screen "Error Counter_2" 320x240
   TextField "Text field_1" at 26,1 size 269x18; Text 'CURRENT SHIFT DATA MINUS 2 (Detil Error)'
   Button "Button_3" at 6,199 size 45x34; TextOff 'Main Page'; PictureOff "Home"
      on Click: ActivateScreen("Main Page", 0)
   Button "Button_1" at 57,206 size 93x28; TextOff 'Back To Data Statistika'; TextOn 'Data Statistika'
      on Click: ActivateScreen("Data Statistika", 0)
   Button "Button_2" at 206,206 size 97x28; TextOff '<----- Back'; TextOn 'Sloft Data'
      on Click: ActivateScreen("Data Time Current Shift_2", 0)
   IOField "I/O field_6" at 6,19 size 132x18; FormatPattern 9999999999999999999999999999999999999999
      ProcessValue <- "DB_DTL1_Cur_ShiftA_2"
   TextField "Text field_9" at 145,21 size 19x15; Text 'S/D'
   IOField "I/O field_7" at 169,20 size 132x18; FormatPattern 9999999999999999999999999999999999999999
      ProcessValue <- "DB_DTL1_Cur_ShiftB_2"
   TextField "Text field_34" at 6,153 size 21x19; Text '6'
   TextField "Text field_33" at 7,133 size 21x19; Text '5'
   TextField "Text field_32" at 7,114 size 21x19; Text '4'
   TextField "Text field_31" at 7,95 size 21x19; Text '3'
   TextField "Text field_30" at 7,76 size 21x19; Text '2'
   TextField "Text field_29" at 7,58 size 21x19; Text '1'
   TextField "Text field_28" at 7,40 size 21x19; Text 'No'
   IOField "I/O field_8" at 225,153 size 26x19; FormatPattern 999
      ProcessValue <- "DB_DTLData_DTL_RS Pneu Er_2.SECOND"
   IOField "I/O field_16" at 200,153 size 25x19; FormatPattern 999
      ProcessValue <- "DB_DTLData_DTL_RS Pneu Er_2.MINUTE"
   IOField "I/O field_17" at 175,153 size 25x19; FormatPattern 999
      ProcessValue <- "DB_DTLData_DTL_RS Pneu Er_2.HOUR"
   TextField "Text field_8" at 29,153 size 145x19; Text 'Reed Swicth Pneumatic Error'
   TextField "Text field_10" at 196,152 size 8x17; Text ':'
   TextField "Text field_21" at 220,153 size 8x17; Text ':'
   IOField "I/O field_21" at 225,94 size 26x19; FormatPattern 999
      ProcessValue <- "Data_DTLData_DTL_Imaje Not In Position[2].SECOND"
   IOField "I/O field_22" at 200,94 size 25x19; FormatPattern 999
      ProcessValue <- "Data_DTLData_DTL_Imaje Not In Position[2].MINUTE"
   IOField "I/O field_23" at 175,94 size 25x19; FormatPattern 999
      ProcessValue <- "Data_DTLData_DTL_Imaje Not In Position[2].HOUR"
   TextField "Text field_25" at 29,95 size 145x19; Text 'Imaje Not In Position'
   IOField "I/O field_18" at 225,76 size 26x19; FormatPattern 999
      ProcessValue <- "Data_DTLData_DTL_Paper R Out[2].SECOND"
   IOField "I/O field_19" at 200,76 size 25x19; FormatPattern 999
      ProcessValue <- "Data_DTLData_DTL_Paper R Out[2].MINUTE"
   IOField "I/O field_20" at 175,76 size 25x19; FormatPattern 999
      ProcessValue <- "Data_DTLData_DTL_Paper R Out[2].HOUR"
   TextField "Text field_22" at 29,76 size 145x19; Text 'Imaje Papper Or Ribbon Out'
   TextField "Text field_2" at 176,43 size 24x15; Text 'Hour'
   IOField "I/O field_10" at 225,134 size 26x19; FormatPattern 999
      ProcessValue <- "DB_DTLData_DTL_Slof Jam_2.SECOND"
   IOField "I/O field_11" at 200,134 size 25x19; FormatPattern 999
      ProcessValue <- "DB_DTLData_DTL_Slof Jam_2.MINUTE"
   IOField "I/O field_12" at 175,134 size 25x19; FormatPattern 999
      ProcessValue <- "DB_DTLData_DTL_Slof Jam_2.HOUR"
   IOField "I/O field_4" at 225,114 size 26x19; FormatPattern 999
      ProcessValue <- "DB_DTLData_DTL_Press Low_2.SECOND"
   IOField "I/O field_5" at 200,114 size 25x19; FormatPattern 999
      ProcessValue <- "DB_DTLData_DTL_Press Low_2.MINUTE"
   IOField "I/O field_9" at 175,114 size 25x19; FormatPattern 999
      ProcessValue <- "DB_DTLData_DTL_Press Low_2.HOUR"
   TextField "Text field_12" at 229,43 size 19x15; Text 'Sec'
   TextField "Text field_11" at 203,43 size 19x15; Text 'Min'
   IOField "I/O field_2" at 225,59 size 26x19; FormatPattern 999
      ProcessValue <- "DB_DTLData_DTL_Imaje Er_2.SECOND"
   IOField "I/O field_1" at 200,59 size 25x19; FormatPattern 999
      ProcessValue <- "DB_DTLData_DTL_Imaje Er_2.MINUTE"
   TextField "Text field_3" at 30,42 size 144x17; Text 'Error Counter'
   TextField "Text field_4" at 29,59 size 145x19; Text 'System Imaje Error'
   TextField "Text field_5" at 29,114 size 145x21; Text 'Pressure Low'
   TextField "Text field_6" at 29,133 size 145x20; Text 'Sloft Jammed'
   IOField "I/O field_3" at 175,59 size 25x19; FormatPattern 999
      ProcessValue <- "DB_DTLData_DTL_Imaje Er_2.HOUR"
   TextField "Text field_13" at 196,58 size 8x17; Text ':'
   TextField "Text field_14" at 196,113 size 8x17; Text ':'
   TextField "Text field_15" at 196,133 size 8x17; Text ':'
   TextField "Text field_17" at 220,58 size 8x17; Text ':'
   TextField "Text field_18" at 220,113 size 8x17; Text ':'
   TextField "Text field_19" at 220,133 size 8x17; Text ':'
   TextField "Text field_23" at 196,75 size 8x17; Text ':'
   TextField "Text field_24" at 220,75 size 8x17; Text ':'
   TextField "Text field_26" at 196,93 size 8x17; Text ':'
   TextField "Text field_27" at 220,93 size 8x17; Text ':'

screen "Error Counter_3" 320x240
   TextField "Text field_1" at 24,1 size 269x18; Text 'CURRENT SHIFT DATA MINUS 3 (Detil Error)'
   Button "Button_3" at 3,198 size 45x34; TextOff 'Main Page'; PictureOff "Home"
      on Click: ActivateScreen("Main Page", 0)
   Button "Button_1" at 54,203 size 93x28; TextOff 'Back To Data Statistika'; TextOn 'Data Statistika'
      on Click: ActivateScreen("Data Statistika", 0)
   Button "Button_2" at 206,203 size 97x28; TextOff '<----- Back'; TextOn 'Sloft Data'
      on Click: ActivateScreen("Data Time Current Shift_3", 0)
   IOField "I/O field_6" at 6,20 size 132x18; FormatPattern 9999999999999999999999999999999999999999
      ProcessValue <- "DB_DTL1_Cur_ShiftA_3"
   TextField "Text field_9" at 145,24 size 19x15; Text 'S/D'
   IOField "I/O field_7" at 169,21 size 132x18; FormatPattern 9999999999999999999999999999999999999999
      ProcessValue <- "DB_DTL1_Cur_ShiftB_3"
   TextField "Text field_34" at 6,153 size 21x19; Text '6'
   TextField "Text field_33" at 7,133 size 21x19; Text '5'
   TextField "Text field_32" at 7,114 size 21x19; Text '4'
   TextField "Text field_31" at 7,95 size 21x19; Text '3'
   TextField "Text field_30" at 7,76 size 21x19; Text '2'
   TextField "Text field_29" at 7,58 size 21x19; Text '1'
   TextField "Text field_28" at 7,40 size 21x19; Text 'No'
   IOField "I/O field_8" at 225,153 size 26x19; FormatPattern 999
      ProcessValue <- "DB_DTLData_DTL_RS Pneu Er_3.SECOND"
   IOField "I/O field_16" at 200,153 size 25x19; FormatPattern 999
      ProcessValue <- "DB_DTLData_DTL_RS Pneu Er_3.MINUTE"
   IOField "I/O field_17" at 175,153 size 25x19; FormatPattern 999
      ProcessValue <- "DB_DTLData_DTL_RS Pneu Er_3.HOUR"
   TextField "Text field_8" at 29,153 size 145x19; Text 'Reed Swicth Pneumatic Error'
   TextField "Text field_10" at 196,152 size 8x17; Text ':'
   TextField "Text field_21" at 220,153 size 8x17; Text ':'
   IOField "I/O field_21" at 225,94 size 26x19; FormatPattern 999
      ProcessValue <- "Data_DTLData_DTL_Imaje Not In Position[3].SECOND"
   IOField "I/O field_22" at 200,94 size 25x19; FormatPattern 999
      ProcessValue <- "Data_DTLData_DTL_Imaje Not In Position[3].MINUTE"
   IOField "I/O field_23" at 175,94 size 25x19; FormatPattern 999
      ProcessValue <- "Data_DTLData_DTL_Imaje Not In Position[3].HOUR"
   TextField "Text field_25" at 29,95 size 145x19; Text 'Imaje Not In Position'
   IOField "I/O field_18" at 225,76 size 26x19; FormatPattern 999
      ProcessValue <- "Data_DTLData_DTL_Paper R Out[3].SECOND"
   IOField "I/O field_19" at 200,76 size 25x19; FormatPattern 999
      ProcessValue <- "Data_DTLData_DTL_Paper R Out[3].MINUTE"
   IOField "I/O field_20" at 175,76 size 25x19; FormatPattern 999
      ProcessValue <- "Data_DTLData_DTL_Paper R Out[3].HOUR"
   TextField "Text field_22" at 29,76 size 145x19; Text 'Imaje Papper Or Ribbon Out'
   TextField "Text field_2" at 176,43 size 24x15; Text 'Hour'
   IOField "I/O field_10" at 225,133 size 26x19; FormatPattern 999
      ProcessValue <- "DB_DTLData_DTL_Slof Jam_3.SECOND"
   IOField "I/O field_11" at 200,133 size 25x19; FormatPattern 999
      ProcessValue <- "DB_DTLData_DTL_Slof Jam_3.MINUTE"
   IOField "I/O field_12" at 175,133 size 25x19; FormatPattern 999
      ProcessValue <- "DB_DTLData_DTL_Slof Jam_3.HOUR"
   IOField "I/O field_4" at 225,114 size 26x19; FormatPattern 999
      ProcessValue <- "DB_DTLData_DTL_Press Low_3.SECOND"
   IOField "I/O field_5" at 200,114 size 25x19; FormatPattern 999
      ProcessValue <- "DB_DTLData_DTL_Press Low_3.MINUTE"
   IOField "I/O field_9" at 175,114 size 25x19; FormatPattern 999
      ProcessValue <- "DB_DTLData_DTL_Press Low_3.HOUR"
   TextField "Text field_12" at 229,43 size 19x15; Text 'Sec'
   TextField "Text field_11" at 203,43 size 19x15; Text 'Min'
   IOField "I/O field_2" at 225,59 size 26x19; FormatPattern 999
      ProcessValue <- "DB_DTLData_DTL_Imaje Er_3.SECOND"
   IOField "I/O field_1" at 200,59 size 25x19; FormatPattern 999
      ProcessValue <- "DB_DTLData_DTL_Imaje Er_3.MINUTE"
   TextField "Text field_3" at 30,42 size 144x17; Text 'Error Counter'
   TextField "Text field_4" at 29,59 size 145x19; Text 'System Imaje Error'
   TextField "Text field_5" at 29,114 size 145x21; Text 'Pressure Low'
   TextField "Text field_6" at 29,133 size 145x20; Text 'Sloft Jammed'
   IOField "I/O field_3" at 175,59 size 25x19; FormatPattern 999
      ProcessValue <- "DB_DTLData_DTL_Imaje Er_3.HOUR"
   TextField "Text field_13" at 196,58 size 8x17; Text ':'
   TextField "Text field_14" at 196,113 size 8x17; Text ':'
   TextField "Text field_15" at 196,132 size 8x17; Text ':'
   TextField "Text field_17" at 220,58 size 8x17; Text ':'
   TextField "Text field_18" at 220,113 size 8x17; Text ':'
   TextField "Text field_19" at 220,132 size 8x17; Text ':'
   TextField "Text field_23" at 196,75 size 8x17; Text ':'
   TextField "Text field_24" at 220,75 size 8x17; Text ':'
   TextField "Text field_26" at 196,93 size 8x17; Text ':'
   TextField "Text field_27" at 220,93 size 8x17; Text ':'

screen "Error Counter_4" 320x240
   TextField "Text field_1" at 25,1 size 269x18; Text 'CURRENT SHIFT DATA MINUS 4 (Detil Error)'
   Button "Button_3" at 0,200 size 45x34; TextOff 'Main Page'; PictureOff "Home"
      on Click: ActivateScreen("Main Page", 0)
   Button "Button_1" at 51,206 size 93x28; TextOff 'Back To Data Statistika'; TextOn 'Data Statistika'
      on Click: ActivateScreen("Data Statistika", 0)
   Button "Button_2" at 207,206 size 97x28; TextOff '<----- Back'; TextOn 'Sloft Data'
      on Click: ActivateScreen("Data Time Current Shift_4", 0)
   IOField "I/O field_6" at 6,20 size 132x18; FormatPattern 9999999999999999999999999999999999999999
      ProcessValue <- "DB_DTL1_Cur_ShiftA_4"
   TextField "Text field_9" at 145,23 size 19x15; Text 'S/D'
   IOField "I/O field_7" at 169,21 size 132x18; FormatPattern 9999999999999999999999999999999999999999
      ProcessValue <- "DB_DTL1_Cur_ShiftB_4"
   TextField "Text field_34" at 6,153 size 21x19; Text '6'
   TextField "Text field_33" at 7,133 size 21x19; Text '5'
   TextField "Text field_32" at 7,114 size 21x19; Text '4'
   TextField "Text field_31" at 7,95 size 21x19; Text '3'
   TextField "Text field_30" at 7,76 size 21x19; Text '2'
   TextField "Text field_29" at 7,58 size 21x19; Text '1'
   TextField "Text field_28" at 7,40 size 21x19; Text 'No'
   IOField "I/O field_8" at 225,153 size 26x19; FormatPattern 999
      ProcessValue <- "DB_DTLData_DTL_RS Pneu Er_4.SECOND"
   IOField "I/O field_16" at 200,153 size 25x19; FormatPattern 999
      ProcessValue <- "DB_DTLData_DTL_RS Pneu Er_4.MINUTE"
   IOField "I/O field_17" at 175,153 size 25x19; FormatPattern 999
      ProcessValue <- "DB_DTLData_DTL_RS Pneu Er_4.HOUR"
   TextField "Text field_8" at 29,153 size 145x19; Text 'Reed Swicth Pneumatic Error'
   TextField "Text field_10" at 196,152 size 8x17; Text ':'
   TextField "Text field_21" at 220,153 size 8x17; Text ':'
   IOField "I/O field_21" at 225,94 size 26x19; FormatPattern 999
      ProcessValue <- "Data_DTLData_DTL_Imaje Not In Position[4].SECOND"
   IOField "I/O field_22" at 200,94 size 25x19; FormatPattern 999
      ProcessValue <- "Data_DTLData_DTL_Imaje Not In Position[4].MINUTE"
   IOField "I/O field_23" at 175,94 size 25x19; FormatPattern 999
      ProcessValue <- "Data_DTLData_DTL_Imaje Not In Position[4].HOUR"
   TextField "Text field_25" at 29,95 size 145x19; Text 'Imaje Not In Position'
   IOField "I/O field_18" at 225,76 size 26x19; FormatPattern 999
      ProcessValue <- "Data_DTLData_DTL_Imaje Not In Position[4].SECOND"
   IOField "I/O field_19" at 200,76 size 25x19; FormatPattern 999
      ProcessValue <- "Data_DTLData_DTL_Paper R Out[4].MINUTE"
   IOField "I/O field_20" at 175,76 size 25x19; FormatPattern 999
      ProcessValue <- "Data_DTLData_DTL_Paper R Out[4].HOUR"
   TextField "Text field_22" at 29,76 size 145x19; Text 'Imaje Papper Or Ribbon Out'
   TextField "Text field_2" at 176,43 size 24x15; Text 'Hour'
   IOField "I/O field_10" at 225,133 size 26x19; FormatPattern 999
      ProcessValue <- "DB_DTLData_DTL_Slof Jam_4.SECOND"
   IOField "I/O field_11" at 200,133 size 25x19; FormatPattern 999
      ProcessValue <- "DB_DTLData_DTL_Slof Jam_4.MINUTE"
   IOField "I/O field_12" at 175,133 size 25x19; FormatPattern 999
      ProcessValue <- "DB_DTLData_DTL_Slof Jam_4.HOUR"
   IOField "I/O field_4" at 225,114 size 26x19; FormatPattern 999
      ProcessValue <- "DB_DTLData_DTL_Press Low_4.SECOND"
   IOField "I/O field_5" at 200,114 size 25x19; FormatPattern 999
      ProcessValue <- "DB_DTLData_DTL_Press Low_4.MINUTE"
   IOField "I/O field_9" at 175,114 size 25x19; FormatPattern 999
      ProcessValue <- "DB_DTLData_DTL_Press Low_4.HOUR"
   TextField "Text field_12" at 229,43 size 19x15; Text 'Sec'
   TextField "Text field_11" at 203,43 size 19x15; Text 'Min'
   IOField "I/O field_2" at 225,59 size 26x19; FormatPattern 999
      ProcessValue <- "DB_DTLData_DTL_Imaje Er_4.SECOND"
   IOField "I/O field_1" at 200,59 size 25x19; FormatPattern 999
      ProcessValue <- "DB_DTLData_DTL_Imaje Er_4.MINUTE"
   TextField "Text field_3" at 30,42 size 144x17; Text 'Error Counter'
   TextField "Text field_4" at 29,59 size 145x19; Text 'System Imaje Error'
   TextField "Text field_5" at 29,114 size 145x21; Text 'Pressure Low'
   TextField "Text field_6" at 29,133 size 145x20; Text 'Sloft Jammed'
   IOField "I/O field_3" at 175,59 size 25x19; FormatPattern 999
      ProcessValue <- "DB_DTLData_DTL_Imaje Er_4.HOUR"
   TextField "Text field_13" at 196,58 size 8x17; Text ':'
   TextField "Text field_14" at 196,113 size 8x17; Text ':'
   TextField "Text field_15" at 196,132 size 8x17; Text ':'
   TextField "Text field_17" at 220,58 size 8x17; Text ':'
   TextField "Text field_18" at 220,113 size 8x17; Text ':'
   TextField "Text field_19" at 220,132 size 8x17; Text ':'
   TextField "Text field_23" at 196,75 size 8x17; Text ':'
   TextField "Text field_24" at 220,75 size 8x17; Text ':'
   TextField "Text field_26" at 196,93 size 8x17; Text ':'
   TextField "Text field_27" at 220,93 size 8x17; Text ':'

screen "Error Counter_5" 320x240
   TextField "Text field_1" at 27,1 size 269x18; Text 'CURRENT SHIFT DATA MINUS 5 (Detil Error)'
   Button "Button_3" at 5,200 size 45x34; TextOff 'Main Page'; PictureOff "Home"
      on Click: ActivateScreen("Main Page", 0)
   Button "Button_1" at 58,206 size 93x28; TextOff 'Back To Data Statistika'; TextOn 'Data Statistika'
      on Click: ActivateScreen("Data Statistika", 0)
   Button "Button_2" at 205,207 size 97x28; TextOff '<----- Back'; TextOn 'Sloft Data'
      on Click: ActivateScreen("Data Time Current Shift_5", 0)
   IOField "I/O field_6" at 6,21 size 132x18; FormatPattern 9999999999999999999999999999999999999999
      ProcessValue <- "DB_DTL1_Cur_ShiftA_5"
   TextField "Text field_9" at 145,23 size 19x15; Text 'S/D'
   IOField "I/O field_7" at 169,21 size 132x18; FormatPattern 9999999999999999999999999999999999999999
      ProcessValue <- "DB_DTL1_Cur_ShiftB_5"
   TextField "Text field_34" at 6,154 size 21x19; Text '6'
   TextField "Text field_33" at 7,134 size 21x19; Text '5'
   TextField "Text field_32" at 7,115 size 21x19; Text '4'
   TextField "Text field_31" at 7,96 size 21x19; Text '3'
   TextField "Text field_30" at 7,77 size 21x19; Text '2'
   TextField "Text field_29" at 7,59 size 21x19; Text '1'
   TextField "Text field_28" at 7,41 size 21x19; Text 'No'
   IOField "I/O field_8" at 225,154 size 26x19; FormatPattern 999
      ProcessValue <- "DB_DTLData_DTL_RS Pneu Er_5.SECOND"
   IOField "I/O field_16" at 200,154 size 25x19; FormatPattern 999
      ProcessValue <- "DB_DTLData_DTL_RS Pneu Er_5.MINUTE"
   IOField "I/O field_17" at 175,154 size 25x19; FormatPattern 999
      ProcessValue <- "DB_DTLData_DTL_RS Pneu Er_5.HOUR"
   TextField "Text field_8" at 29,154 size 145x19; Text 'Reed Swicth Pneumatic Error'
   TextField "Text field_10" at 196,153 size 8x17; Text ':'
   TextField "Text field_21" at 220,154 size 8x17; Text ':'
   IOField "I/O field_21" at 225,95 size 26x19; FormatPattern 999
      ProcessValue <- "Data_DTLData_DTL_Imaje Not In Position[5].SECOND"
   IOField "I/O field_22" at 200,95 size 25x19; FormatPattern 999
      ProcessValue <- "Data_DTLData_DTL_Imaje Not In Position[5].MINUTE"
   IOField "I/O field_23" at 175,95 size 25x19; FormatPattern 999
      ProcessValue <- "Data_DTLData_DTL_Imaje Not In Position[5].HOUR"
   TextField "Text field_25" at 29,96 size 145x19; Text 'Imaje Not In Position'
   IOField "I/O field_18" at 225,77 size 26x19; FormatPattern 999
      ProcessValue <- "Data_DTLData_DTL_Paper R Out[5].SECOND"
   IOField "I/O field_19" at 200,77 size 25x19; FormatPattern 999
      ProcessValue <- "Data_DTLData_DTL_Paper R Out[5].MINUTE"
   IOField "I/O field_20" at 175,77 size 25x19; FormatPattern 999
      ProcessValue <- "Data_DTLData_DTL_Paper R Out[5].HOUR"
   TextField "Text field_22" at 29,77 size 145x19; Text 'Imaje Papper Or Ribbon Out'
   TextField "Text field_2" at 176,44 size 24x15; Text 'Hour'
   IOField "I/O field_10" at 225,134 size 26x19; FormatPattern 999
      ProcessValue <- "DB_DTLData_DTL_Slof Jam_5.SECOND"
   IOField "I/O field_11" at 200,134 size 25x19; FormatPattern 999
      ProcessValue <- "DB_DTLData_DTL_Slof Jam_5.MINUTE"
   IOField "I/O field_12" at 175,134 size 25x19; FormatPattern 999
      ProcessValue <- "DB_DTLData_DTL_Slof Jam_5.HOUR"
   IOField "I/O field_4" at 225,115 size 26x19; FormatPattern 999
      ProcessValue <- "DB_DTLData_DTL_Press Low_5.SECOND"
   IOField "I/O field_5" at 200,115 size 25x19; FormatPattern 999
      ProcessValue <- "DB_DTLData_DTL_Press Low_5.MINUTE"
   IOField "I/O field_9" at 175,115 size 25x19; FormatPattern 999
      ProcessValue <- "DB_DTLData_DTL_Press Low_5.HOUR"
   TextField "Text field_12" at 229,44 size 19x15; Text 'Sec'
   TextField "Text field_11" at 203,44 size 19x15; Text 'Min'
   IOField "I/O field_2" at 225,60 size 26x19; FormatPattern 999
      ProcessValue <- "DB_DTLData_DTL_Imaje Er_5.SECOND"
   IOField "I/O field_1" at 200,60 size 25x19; FormatPattern 999
      ProcessValue <- "DB_DTLData_DTL_Imaje Er_5.MINUTE"
   TextField "Text field_3" at 30,43 size 144x17; Text 'Error Counter'
   TextField "Text field_4" at 29,60 size 145x19; Text 'System Imaje Error'
   TextField "Text field_5" at 29,115 size 145x21; Text 'Pressure Low'
   TextField "Text field_6" at 29,134 size 145x20; Text 'Sloft Jammed'
   IOField "I/O field_3" at 175,60 size 25x19; FormatPattern 999
      ProcessValue <- "DB_DTLData_DTL_Imaje Er_5.HOUR"
   TextField "Text field_13" at 196,59 size 8x17; Text ':'
   TextField "Text field_14" at 196,114 size 8x17; Text ':'
   TextField "Text field_15" at 196,133 size 8x17; Text ':'
   TextField "Text field_17" at 220,59 size 8x17; Text ':'
   TextField "Text field_18" at 220,114 size 8x17; Text ':'
   TextField "Text field_19" at 220,133 size 8x17; Text ':'
   TextField "Text field_23" at 196,76 size 8x17; Text ':'
   TextField "Text field_24" at 220,76 size 8x17; Text ':'
   TextField "Text field_26" at 196,94 size 8x17; Text ':'
   TextField "Text field_27" at 220,94 size 8x17; Text ':'

screen "Statistik Parameter" 320x240
   TextField "Text field_13" at 186,102 size 26x12; Text 'Hour'
   TextField "Text field_17" at 122,102 size 34x12; Text 'Second'
   TextField "Text field_10" at 118,88 size 86x16; Text 'Time Shift Setting'
   TextField "Text field_4" at 71,19 size 47x13; Text 'Day (1-31)'
   TextField "Text field_6" at 196,19 size 21x13; Text 'Year'
   TextField "Text field_5" at 119,19 size 61x12; Text 'Month (1-12)'
   TextField "Text field_1" at 6,1 size 143x17; Text 'STATISTIKA PARAMETER'
   TextField "Text field_2" at 9,32 size 62x15; Text 'Date Setting'
   TextField "Text field_3" at 10,65 size 61x15; Text 'Time Setting'
   TextField "Text field_7" at 67,54 size 52x12; Text 'Hour (0-23)'
   TextField "Text field_8" at 119,53 size 59x12; Text 'Minute (0-59)'
   TextField "Text field_9" at 176,53 size 64x12; Text 'Second (0-59)'
   IOField "I/O field_6" at 72,33 size 42x20; FormatPattern 99
      ProcessValue <- "DB_Integer_IDay"
   Button "Button_1" at 256,50 size 57x23; TextOff 'Execute'; TextOn 'OK'
      on Release: ResetBit("DB_Bool1_F_Set Time Day")
      on Press: SetBit("DB_Bool1_F_Set Time Day")
   TextField "Text field_11" at 11,117 size 33x15; Text 'Shift 1'
   TextField "Text field_15" at 49,102 size 26x12; Text 'Hour'
   TextField "Text field_16" at 85,102 size 30x12; Text 'Minute'
   IOField "I/O field_7" at 81,115 size 35x20; FormatPattern 99
      ProcessValue <- "DB_Integer_S1AMinute"
   IOField "I/O field_8" at 119,115 size 35x20; FormatPattern 99
      ProcessValue <- "DB_Integer_S1ASecond"
   TextField "Text field_12" at 160,114 size 17x15; Text 's/d'
   IOField "I/O field_9" at 180,115 size 35x20; FormatPattern 99
      ProcessValue <- "DB_Integer_S1BHour"
   TextField "Text field_14" at 221,102 size 30x12; Text 'Minute'
   TextField "Text field_18" at 256,102 size 34x12; Text 'Second'
   IOField "I/O field_11" at 218,115 size 35x20; FormatPattern 99
      ProcessValue <- "DB_Integer_S1BMinute"
   IOField "I/O field_12" at 256,115 size 35x20; FormatPattern 99
      ProcessValue <- "DB_Integer_S1BSecond"
   TextField "Text field_19" at 10,141 size 33x15; Text 'Shift 2'
   IOField "I/O field_13" at 43,139 size 35x20; FormatPattern 99
      ProcessValue <- "DB_Integer_S2AHour"
   IOField "I/O field_14" at 81,139 size 35x20; FormatPattern 99
      ProcessValue <- "DB_Integer_S2AMinute"
   IOField "I/O field_15" at 119,139 size 35x20; FormatPattern 99
      ProcessValue <- "DB_Integer_S2ASecond"
   TextField "Text field_23" at 160,140 size 17x15; Text 's/d'
   IOField "I/O field_16" at 180,139 size 35x20; FormatPattern 99
      ProcessValue <- "DB_Integer_S2BHour"
   IOField "I/O field_17" at 218,139 size 35x20; FormatPattern 99
      ProcessValue <- "DB_Integer_S2BMinute"
   IOField "I/O field_18" at 256,139 size 35x20; FormatPattern 99
      ProcessValue <- "DB_Integer_S2BSecond"
   TextField "Text field_27" at 9,165 size 33x15; Text 'Shift 3'
   IOField "I/O field_19" at 43,163 size 35x20; FormatPattern 99
      ProcessValue <- "DB_Integer_S3AHour"
   IOField "I/O field_20" at 81,163 size 35x20; FormatPattern 99
      ProcessValue <- "DB_Integer_S3AMinute"
   IOField "I/O field_21" at 119,163 size 35x20; FormatPattern 99
      ProcessValue <- "DB_Integer_S3ASecond"
   TextField "Text field_31" at 160,164 size 17x15; Text 's/d'
   IOField "I/O field_22" at 180,163 size 35x20; FormatPattern 99
      ProcessValue <- "DB_Integer_S3BHour"
   IOField "I/O field_23" at 218,163 size 35x20; FormatPattern 99
      ProcessValue <- "DB_Integer_S3BMinute"
   IOField "I/O field_24" at 256,163 size 35x20; FormatPattern 99
      ProcessValue <- "DB_Integer_S3BSecond"
   IOField "I/O field_10" at 43,115 size 35x20; FormatPattern 99
      ProcessValue <- "DB_Integer_S1AHour"
   IOField "I/O field_1" at 125,33 size 43x20; FormatPattern 99
      ProcessValue <- "DB_Integer_IMonth"
   IOField "I/O field_2" at 180,33 size 52x20; FormatPattern 9999
      ProcessValue <- "DB_Integer_IYear"
   IOField "I/O field_3" at 72,66 size 40x20; FormatPattern 99
      ProcessValue <- "DB_Integer_IHour"
   IOField "I/O field_4" at 129,66 size 40x20; FormatPattern 99
      ProcessValue <- "DB_Integer_IMinute"
   IOField "I/O field_5" at 185,66 size 40x20; FormatPattern 99
      ProcessValue <- "DB_Integer_ISecond"
   IOField "I/O field_25" at 163,1 size 155x23; FormatPattern 9999999999999999999999999999999999999999
      ProcessValue <- "DB_DTL1_Output"
   Button "Button_2" at 138,185 size 57x24; TextOff 'Execute'; TextOn 'OK'
   Button "Button_4" at 3,211 size 35x27; TextOff 'Main Page'; PictureOff "Home"
      on Click: ActivateScreen("Main Page", 0)

screen "Data Time Current Shift" 320x240
   IOField "I/O field_12" at 252,92 size 56x19; FormatPattern 999.99; Unit   %
      ProcessValue <- "Data_Real_%Mesin Run Baypass[0]"
   IOField "I/O field_13" at 252,110 size 56x21; FormatPattern 999.99; Unit   %
      ProcessValue <- "Data_Real_%Mesin Stop[0]"
   IOField "I/O field_14" at 252,130 size 56x20; FormatPattern 999.99; Unit   %
      ProcessValue <- "Data_Real_%Mesin Error[0]"
   IOField "I/O field_11" at 252,75 size 56x18; FormatPattern 999.99; Unit   %
      ProcessValue <- "Data_Real_%Mesin Run[0]"
   Button "Button_1" at 43,206 size 90x32; TextOff 'Back To Statistika Data'; TextOn 'Statistika Data'
      on Click: ActivateScreen("Data Statistika", 0)
   Button "Button_3" at 0,204 size 41x34; TextOff 'Main Page'; PictureOff "Home"
      on Click: ActivateScreen("Main Page", 0)
   Button "Button_2" at 236,207 size 80x30; TextOff 'Next Data --->'; TextOn 'Detail Error'
      on Click: ActivateScreen("Error Counter", 0)
   TextField "Text field_1" at 92,0 size 174x18; Text 'CURRENT SHIFT (Time Data)'
   IOField "I/O field_6" at 7,24 size 132x18; FormatPattern 9999999999999999999999999999999999999999
      ProcessValue <- "DB_DTL1_Cur_ShiftA"
   TextField "Text field_9" at 145,23 size 19x15; Text 'S/D'
   IOField "I/O field_7" at 170,24 size 132x18; FormatPattern 9999999999999999999999999999999999999999
      ProcessValue <- "DB_DTL1_Cur_ShiftB"
   TextField "Text field_32" at 7,130 size 21x19; Text '4'
   TextField "Text field_31" at 7,111 size 21x19; Text '3'
   TextField "Text field_30" at 7,92 size 21x19; Text '2'
   TextField "Text field_29" at 7,74 size 21x19; Text '1'
   TextField "Text field_28" at 7,56 size 21x19; Text 'No'
   IOField "I/O field_21" at 225,110 size 26x19; FormatPattern 999
      ProcessValue <- "Data_DTLData_DTL_Mesin Stop[0].SECOND"
   IOField "I/O field_22" at 200,110 size 25x19; FormatPattern 999
      ProcessValue <- "Data_DTLData_DTL_Mesin Stop[0].MINUTE"
   IOField "I/O field_23" at 175,110 size 25x19; FormatPattern 999
      ProcessValue <- "Data_DTLData_DTL_Mesin Stop[0].HOUR"
   TextField "Text field_25" at 29,111 size 145x19; Text 'Stop'
   IOField "I/O field_18" at 225,92 size 26x19; FormatPattern 999
      ProcessValue <- "Data_DTLData_DTL_Mesin Run Baypass[0].SECOND"
   IOField "I/O field_19" at 200,92 size 25x19; FormatPattern 999
      ProcessValue <- "Data_DTLData_DTL_Mesin Run Baypass[0].MINUTE"
   IOField "I/O field_20" at 175,92 size 25x19; FormatPattern 999
      ProcessValue <- "Data_DTLData_DTL_Mesin Run Baypass[0].HOUR"
   TextField "Text field_22" at 29,92 size 145x19; Text 'Running Bypass Stamp'
   TextField "Text field_2" at 176,59 size 24x15; Text 'Hour'
   IOField "I/O field_4" at 225,130 size 26x19; FormatPattern 999
      ProcessValue <- "Data_DTLData_DTL_Mesin Error[0].SECOND"
   IOField "I/O field_5" at 200,130 size 25x19; FormatPattern 999
      ProcessValue <- "Data_DTLData_DTL_Mesin Error[0].MINUTE"
   IOField "I/O field_9" at 175,130 size 25x19; FormatPattern 999
      ProcessValue <- "Data_DTLData_DTL_Mesin Error[0].HOUR"
   TextField "Text field_12" at 229,59 size 19x15; Text 'Sec'
   TextField "Text field_11" at 203,59 size 19x15; Text 'Min'
   IOField "I/O field_2" at 225,75 size 26x19; FormatPattern 999
      ProcessValue <- "Data_DTLData_DTL_Mesin Run[0].SECOND"
   IOField "I/O field_3" at 200,75 size 25x19; FormatPattern 999
      ProcessValue <- "Data_DTLData_DTL_Mesin Run[0].MINUTE"
   TextField "Text field_3" at 30,58 size 144x17; Text 'Time Counter Machine'
   TextField "Text field_4" at 29,75 size 145x19; Text 'Running'
   TextField "Text field_5" at 29,130 size 145x20; Text 'Error'
   IOField "I/O field_24" at 175,75 size 25x19; FormatPattern 999
      ProcessValue <- "Data_DTLData_DTL_Mesin Run[0].HOUR"
   TextField "Text field_13" at 196,74 size 8x17; Text ':'
   TextField "Text field_14" at 196,129 size 8x17; Text ':'
   TextField "Text field_17" at 220,74 size 8x17; Text ':'
   TextField "Text field_18" at 220,129 size 8x17; Text ':'
   TextField "Text field_23" at 196,91 size 8x17; Text ':'
   TextField "Text field_24" at 220,91 size 8x17; Text ':'
   TextField "Text field_26" at 196,109 size 8x17; Text ':'
   TextField "Text field_27" at 220,109 size 8x17; Text ':'
   Button "Button_4" at 146,207 size 87x30; TextOff '<--- Back Data'; TextOn 'Sloft Data'
      on Click: ActivateScreen("Data Current Shift", 0)

screen "Data Time Current Shift_1" 320x240
   IOField "I/O field_12" at 252,92 size 56x19; FormatPattern 999.99; Unit   %
      ProcessValue <- "Data_Real_%Mesin Run Baypass[1]"
   IOField "I/O field_13" at 252,110 size 56x21; FormatPattern 999.99; Unit   %
      ProcessValue <- "Data_Real_%Mesin Stop[1]"
   IOField "I/O field_14" at 252,130 size 56x20; FormatPattern 999.99; Unit   %
      ProcessValue <- "Data_Real_%Mesin Error[1]"
   IOField "I/O field_11" at 252,75 size 56x18; FormatPattern 999.99; Unit   %
      ProcessValue <- "Data_Real_%Mesin Run[1]"
   Button "Button_1" at 47,206 size 90x32; TextOff 'Back To Statistika Data'; TextOn 'Statistika Data'
      on Click: ActivateScreen("Data Statistika", 0)
   Button "Button_3" at 1,205 size 41x34; TextOff 'Main Page'; PictureOff "Home"
      on Click: ActivateScreen("Main Page", 0)
   TextField "Text field_1" at 47,0 size 230x18; Text 'CURRENT SHIFT MINUS 1 (Time Data)'
   IOField "I/O field_6" at 7,24 size 132x18; FormatPattern 9999999999999999999999999999999999999999
      ProcessValue <- "DB_DTL1_Cur_ShiftA_1"
   TextField "Text field_9" at 145,23 size 19x15; Text 'S/D'
   IOField "I/O field_7" at 170,24 size 132x18; FormatPattern 9999999999999999999999999999999999999999
      ProcessValue <- "DB_DTL1_Cur_ShiftB_1"
   TextField "Text field_32" at 7,130 size 21x19; Text '4'
   TextField "Text field_31" at 7,111 size 21x19; Text '3'
   TextField "Text field_30" at 7,92 size 21x19; Text '2'
   TextField "Text field_29" at 7,74 size 21x19; Text '1'
   TextField "Text field_28" at 7,56 size 21x19; Text 'No'
   IOField "I/O field_21" at 225,110 size 26x19; FormatPattern 999
      ProcessValue <- "Data_DTLData_DTL_Mesin Stop[1].SECOND"
   IOField "I/O field_22" at 200,110 size 25x19; FormatPattern 999
      ProcessValue <- "Data_DTLData_DTL_Mesin Stop[1].MINUTE"
   IOField "I/O field_23" at 175,110 size 25x19; FormatPattern 999
      ProcessValue <- "Data_DTLData_DTL_Mesin Stop[1].HOUR"
   TextField "Text field_25" at 29,111 size 145x19; Text 'Stop'
   IOField "I/O field_18" at 225,92 size 26x19; FormatPattern 999
      ProcessValue <- "Data_DTLData_DTL_Mesin Run Baypass[1].SECOND"
   IOField "I/O field_19" at 200,92 size 25x19; FormatPattern 999
      ProcessValue <- "Data_DTLData_DTL_Mesin Run Baypass[1].MINUTE"
   IOField "I/O field_20" at 175,92 size 25x19; FormatPattern 999
      ProcessValue <- "Data_DTLData_DTL_Mesin Run Baypass[1].HOUR"
   TextField "Text field_22" at 29,92 size 145x19; Text 'Running Bypass Stamp'
   TextField "Text field_2" at 176,59 size 24x15; Text 'Hour'
   IOField "I/O field_4" at 225,130 size 26x19; FormatPattern 999
      ProcessValue <- "Data_DTLData_DTL_Mesin Error[1].SECOND"
   IOField "I/O field_5" at 200,130 size 25x19; FormatPattern 999
      ProcessValue <- "Data_DTLData_DTL_Mesin Error[1].MINUTE"
   IOField "I/O field_9" at 175,130 size 25x19; FormatPattern 999
      ProcessValue <- "Data_DTLData_DTL_Mesin Error[1].HOUR"
   TextField "Text field_12" at 229,59 size 19x15; Text 'Sec'
   TextField "Text field_11" at 203,59 size 19x15; Text 'Min'
   IOField "I/O field_2" at 225,75 size 26x19; FormatPattern 999
      ProcessValue <- "Data_DTLData_DTL_Mesin Run[1].SECOND"
   IOField "I/O field_3" at 200,75 size 25x19; FormatPattern 999
      ProcessValue <- "Data_DTLData_DTL_Mesin Run[1].MINUTE"
   TextField "Text field_3" at 30,58 size 144x17; Text 'Time Counter Machine'
   TextField "Text field_4" at 29,75 size 145x19; Text 'Running'
   TextField "Text field_5" at 29,130 size 145x20; Text 'Error'
   IOField "I/O field_24" at 175,75 size 25x19; FormatPattern 999
      ProcessValue <- "Data_DTLData_DTL_Mesin Run[1].HOUR"
   TextField "Text field_13" at 196,74 size 8x17; Text ':'
   TextField "Text field_14" at 196,129 size 8x17; Text ':'
   TextField "Text field_17" at 220,74 size 8x17; Text ':'
   TextField "Text field_18" at 220,129 size 8x17; Text ':'
   TextField "Text field_23" at 196,91 size 8x17; Text ':'
   TextField "Text field_24" at 220,91 size 8x17; Text ':'
   TextField "Text field_26" at 196,109 size 8x17; Text ':'
   TextField "Text field_27" at 220,109 size 8x17; Text ':'
   Button "Button_2" at 236,207 size 80x30; TextOff 'Next Data --->'; TextOn 'Detail Error'
      on Click: ActivateScreen("Error Counter_1", 0)
   Button "Button_4" at 146,207 size 87x30; TextOff '<--- Back Data'; TextOn 'Sloft Data'
      on Click: ActivateScreen("Data Current Shift_1", 0)

screen "Data Time Current Shift_2" 320x240
   IOField "I/O field_12" at 252,92 size 56x19; FormatPattern 999.99; Unit   %
      ProcessValue <- "Data_Real_%Mesin Run Baypass[2]"
   IOField "I/O field_13" at 252,110 size 56x21; FormatPattern 999.99; Unit   %
      ProcessValue <- "Data_Real_%Mesin Stop[2]"
   IOField "I/O field_14" at 252,130 size 56x20; FormatPattern 999.99; Unit   %
      ProcessValue <- "Data_Real_%Mesin Error[2]"
   IOField "I/O field_11" at 252,75 size 56x18; FormatPattern 999.99; Unit   %
      ProcessValue <- "Data_Real_%Mesin Run[2]"
   IOField "I/O field_6" at 7,24 size 132x18; FormatPattern 9999999999999999999999999999999999999999
      ProcessValue <- "DB_DTL1_Cur_ShiftA_2"
   TextField "Text field_9" at 145,23 size 19x15; Text 'S/D'
   IOField "I/O field_7" at 170,24 size 132x18; FormatPattern 9999999999999999999999999999999999999999
      ProcessValue <- "DB_DTL1_Cur_ShiftB_2"
   TextField "Text field_32" at 7,130 size 21x19; Text '4'
   TextField "Text field_31" at 7,111 size 21x19; Text '3'
   TextField "Text field_30" at 7,92 size 21x19; Text '2'
   TextField "Text field_29" at 7,74 size 21x19; Text '1'
   TextField "Text field_28" at 7,56 size 21x19; Text 'No'
   IOField "I/O field_21" at 225,110 size 26x19; FormatPattern 999
      ProcessValue <- "Data_DTLData_DTL_Mesin Stop[2].SECOND"
   IOField "I/O field_22" at 200,110 size 25x19; FormatPattern 999
      ProcessValue <- "Data_DTLData_DTL_Mesin Stop[2].MINUTE"
   IOField "I/O field_23" at 175,110 size 25x19; FormatPattern 999
      ProcessValue <- "Data_DTLData_DTL_Mesin Stop[2].HOUR"
   TextField "Text field_25" at 29,111 size 145x19; Text 'Stop'
   IOField "I/O field_18" at 225,92 size 26x19; FormatPattern 999
      ProcessValue <- "Data_DTLData_DTL_Mesin Run Baypass[2].SECOND"
   IOField "I/O field_19" at 200,92 size 25x19; FormatPattern 999
      ProcessValue <- "Data_DTLData_DTL_Mesin Run Baypass[2].MINUTE"
   IOField "I/O field_20" at 175,92 size 25x19; FormatPattern 999
      ProcessValue <- "Data_DTLData_DTL_Mesin Run Baypass[2].HOUR"
   TextField "Text field_22" at 29,92 size 145x19; Text 'Running Bypass Stamp'
   TextField "Text field_2" at 176,59 size 24x15; Text 'Hour'
   IOField "I/O field_4" at 225,130 size 26x19; FormatPattern 999
      ProcessValue <- "Data_DTLData_DTL_Mesin Error[2].SECOND"
   IOField "I/O field_5" at 200,130 size 25x19; FormatPattern 999
      ProcessValue <- "Data_DTLData_DTL_Mesin Error[2].MINUTE"
   IOField "I/O field_9" at 175,130 size 25x19; FormatPattern 999
      ProcessValue <- "Data_DTLData_DTL_Mesin Error[2].HOUR"
   TextField "Text field_12" at 229,59 size 19x15; Text 'Sec'
   TextField "Text field_11" at 203,59 size 19x15; Text 'Min'
   IOField "I/O field_2" at 225,75 size 26x19; FormatPattern 999
      ProcessValue <- "Data_DTLData_DTL_Mesin Run[2].SECOND"
   IOField "I/O field_3" at 200,75 size 25x19; FormatPattern 999
      ProcessValue <- "Data_DTLData_DTL_Mesin Run[2].MINUTE"
   TextField "Text field_3" at 30,58 size 144x17; Text 'Time Counter Machine'
   TextField "Text field_4" at 29,75 size 145x19; Text 'Running'
   TextField "Text field_5" at 29,130 size 145x20; Text 'Error'
   IOField "I/O field_24" at 175,75 size 25x19; FormatPattern 999
      ProcessValue <- "Data_DTLData_DTL_Mesin Run[2].HOUR"
   TextField "Text field_13" at 196,74 size 8x17; Text ':'
   TextField "Text field_14" at 196,129 size 8x17; Text ':'
   TextField "Text field_17" at 220,74 size 8x17; Text ':'
   TextField "Text field_18" at 220,129 size 8x17; Text ':'
   TextField "Text field_23" at 196,91 size 8x17; Text ':'
   TextField "Text field_24" at 220,91 size 8x17; Text ':'
   TextField "Text field_26" at 196,109 size 8x17; Text ':'
   TextField "Text field_27" at 220,109 size 8x17; Text ':'
   Button "Button_1" at 47,206 size 90x32; TextOff 'Back To Statistika Data'; TextOn 'Statistika Data'
      on Click: ActivateScreen("Data Statistika", 0)
   Button "Button_3" at 1,205 size 41x34; TextOff 'Main Page'; PictureOff "Home"
      on Click: ActivateScreen("Main Page", 0)
   Button "Button_2" at 236,207 size 80x30; TextOff 'Next Data --->'; TextOn 'Detail Error'
      on Click: ActivateScreen("Error Counter_2", 0)
   Button "Button_4" at 146,207 size 87x30; TextOff '<--- Back Data'; TextOn 'Sloft Data'
      on Click: ActivateScreen("Data Current Shift_2", 0)
   TextField "Text field_1" at 47,0 size 230x18; Text 'CURRENT SHIFT MINUS 2 (Time Data)'

screen "Data Time Current Shift_3" 320x240
   IOField "I/O field_12" at 252,92 size 56x19; FormatPattern 999.99; Unit   %
      ProcessValue <- "Data_Real_%Mesin Run Baypass[3]"
   IOField "I/O field_13" at 252,110 size 56x21; FormatPattern 999.99; Unit   %
      ProcessValue <- "Data_Real_%Mesin Stop[3]"
   IOField "I/O field_14" at 252,130 size 56x20; FormatPattern 999.99; Unit   %
      ProcessValue <- "Data_Real_%Mesin Error[3]"
   IOField "I/O field_11" at 252,75 size 56x18; FormatPattern 999.99; Unit   %
      ProcessValue <- "Data_Real_%Mesin Run[3]"
   IOField "I/O field_6" at 7,24 size 132x18; FormatPattern 9999999999999999999999999999999999999999
      ProcessValue <- "DB_DTL1_Cur_ShiftA_3"
   TextField "Text field_9" at 145,23 size 19x15; Text 'S/D'
   IOField "I/O field_7" at 170,24 size 132x18; FormatPattern 9999999999999999999999999999999999999999
      ProcessValue <- "DB_DTL1_Cur_ShiftB_3"
   TextField "Text field_32" at 7,130 size 21x19; Text '4'
   TextField "Text field_31" at 7,111 size 21x19; Text '3'
   TextField "Text field_30" at 7,92 size 21x19; Text '2'
   TextField "Text field_29" at 7,74 size 21x19; Text '1'
   TextField "Text field_28" at 7,56 size 21x19; Text 'No'
   IOField "I/O field_21" at 225,110 size 26x19; FormatPattern 999
      ProcessValue <- "Data_DTLData_DTL_Mesin Stop[3].SECOND"
   IOField "I/O field_22" at 200,110 size 25x19; FormatPattern 999
      ProcessValue <- "Data_DTLData_DTL_Mesin Stop[3].MINUTE"
   IOField "I/O field_23" at 175,110 size 25x19; FormatPattern 999
      ProcessValue <- "Data_DTLData_DTL_Mesin Stop[3].HOUR"
   TextField "Text field_25" at 29,111 size 145x19; Text 'Stop'
   IOField "I/O field_18" at 225,92 size 26x19; FormatPattern 999
      ProcessValue <- "Data_DTLData_DTL_Mesin Run Baypass[3].SECOND"
   IOField "I/O field_19" at 200,92 size 25x19; FormatPattern 999
      ProcessValue <- "Data_DTLData_DTL_Mesin Run Baypass[3].MINUTE"
   IOField "I/O field_20" at 175,92 size 25x19; FormatPattern 999
      ProcessValue <- "Data_DTLData_DTL_Mesin Run Baypass[3].HOUR"
   TextField "Text field_22" at 29,92 size 145x19; Text 'Running Bypass Stamp'
   TextField "Text field_2" at 176,59 size 24x15; Text 'Hour'
   IOField "I/O field_4" at 225,130 size 26x19; FormatPattern 999
      ProcessValue <- "Data_DTLData_DTL_Mesin Error[3].SECOND"
   IOField "I/O field_5" at 200,130 size 25x19; FormatPattern 999
      ProcessValue <- "Data_DTLData_DTL_Mesin Error[3].MINUTE"
   IOField "I/O field_9" at 175,130 size 25x19; FormatPattern 999
      ProcessValue <- "Data_DTLData_DTL_Mesin Error[3].HOUR"
   TextField "Text field_12" at 229,59 size 19x15; Text 'Sec'
   TextField "Text field_11" at 203,59 size 19x15; Text 'Min'
   IOField "I/O field_2" at 225,75 size 26x19; FormatPattern 999
      ProcessValue <- "Data_DTLData_DTL_Mesin Run[3].SECOND"
   IOField "I/O field_3" at 200,75 size 25x19; FormatPattern 999
      ProcessValue <- "Data_DTLData_DTL_Mesin Run[3].MINUTE"
   TextField "Text field_3" at 30,58 size 144x17; Text 'Time Counter Machine'
   TextField "Text field_4" at 29,75 size 145x19; Text 'Running'
   TextField "Text field_5" at 29,130 size 145x20; Text 'Error'
   IOField "I/O field_24" at 175,75 size 25x19; FormatPattern 999
      ProcessValue <- "Data_DTLData_DTL_Mesin Run[3].HOUR"
   TextField "Text field_13" at 196,74 size 8x17; Text ':'
   TextField "Text field_14" at 196,129 size 8x17; Text ':'
   TextField "Text field_17" at 220,74 size 8x17; Text ':'
   TextField "Text field_18" at 220,129 size 8x17; Text ':'
   TextField "Text field_23" at 196,91 size 8x17; Text ':'
   TextField "Text field_24" at 220,91 size 8x17; Text ':'
   TextField "Text field_26" at 196,109 size 8x17; Text ':'
   TextField "Text field_27" at 220,109 size 8x17; Text ':'
   Button "Button_1" at 47,206 size 90x32; TextOff 'Back To Statistika Data'; TextOn 'Statistika Data'
      on Click: ActivateScreen("Data Statistika", 0)
   Button "Button_3" at 1,205 size 41x34; TextOff 'Main Page'; PictureOff "Home"
      on Click: ActivateScreen("Main Page", 0)
   Button "Button_2" at 236,207 size 80x30; TextOff 'Next Data --->'; TextOn 'Detail Error'
      on Click: ActivateScreen("Error Counter_3", 0)
   Button "Button_4" at 146,207 size 87x30; TextOff '<--- Back Data'; TextOn 'Sloft Data'
      on Click: ActivateScreen("Data Current Shift_3", 0)
   TextField "Text field_1" at 47,0 size 230x18; Text 'CURRENT SHIFT MINUS 3 (Time Data)'

screen "Data Time Current Shift_4" 320x240
   IOField "I/O field_12" at 252,92 size 56x19; FormatPattern 999.99; Unit   %
      ProcessValue <- "Data_Real_%Mesin Run Baypass[4]"
   IOField "I/O field_13" at 252,110 size 56x21; FormatPattern 999.99; Unit   %
      ProcessValue <- "Data_Real_%Mesin Stop[4]"
   IOField "I/O field_14" at 252,130 size 56x20; FormatPattern 999.99; Unit   %
      ProcessValue <- "Data_Real_%Mesin Error[4]"
   IOField "I/O field_11" at 252,75 size 56x18; FormatPattern 999.99; Unit   %
      ProcessValue <- "Data_Real_%Mesin Run[4]"
   IOField "I/O field_6" at 7,24 size 132x18; FormatPattern 9999999999999999999999999999999999999999
      ProcessValue <- "DB_DTL1_Cur_ShiftA_4"
   TextField "Text field_9" at 145,23 size 19x15; Text 'S/D'
   IOField "I/O field_7" at 170,24 size 132x18; FormatPattern 9999999999999999999999999999999999999999
      ProcessValue <- "DB_DTL1_Cur_ShiftB_4"
   TextField "Text field_32" at 7,130 size 21x19; Text '4'
   TextField "Text field_31" at 7,111 size 21x19; Text '3'
   TextField "Text field_30" at 7,92 size 21x19; Text '2'
   TextField "Text field_29" at 7,74 size 21x19; Text '1'
   TextField "Text field_28" at 7,56 size 21x19; Text 'No'
   IOField "I/O field_21" at 225,110 size 26x19; FormatPattern 999
      ProcessValue <- "Data_DTLData_DTL_Mesin Stop[4].SECOND"
   IOField "I/O field_22" at 200,110 size 25x19; FormatPattern 999
      ProcessValue <- "Data_DTLData_DTL_Mesin Stop[4].MINUTE"
   IOField "I/O field_23" at 175,110 size 25x19; FormatPattern 999
      ProcessValue <- "Data_DTLData_DTL_Mesin Stop[4].HOUR"
   TextField "Text field_25" at 29,111 size 145x19; Text 'Stop'
   IOField "I/O field_18" at 225,92 size 26x19; FormatPattern 999
      ProcessValue <- "Data_DTLData_DTL_Mesin Run Baypass[4].SECOND"
   IOField "I/O field_19" at 200,92 size 25x19; FormatPattern 999
      ProcessValue <- "Data_DTLData_DTL_Mesin Run Baypass[4].MINUTE"
   IOField "I/O field_20" at 175,92 size 25x19; FormatPattern 999
      ProcessValue <- "Data_DTLData_DTL_Mesin Run Baypass[4].HOUR"
   TextField "Text field_22" at 29,92 size 145x19; Text 'Running Bypass Stamp'
   TextField "Text field_2" at 176,59 size 24x15; Text 'Hour'
   IOField "I/O field_4" at 225,130 size 26x19; FormatPattern 999
      ProcessValue <- "Data_DTLData_DTL_Mesin Error[4].SECOND"
   IOField "I/O field_5" at 200,130 size 25x19; FormatPattern 999
      ProcessValue <- "Data_DTLData_DTL_Mesin Error[4].MINUTE"
   IOField "I/O field_9" at 175,130 size 25x19; FormatPattern 999
      ProcessValue <- "Data_DTLData_DTL_Mesin Error[4].HOUR"
   TextField "Text field_12" at 229,59 size 19x15; Text 'Sec'
   TextField "Text field_11" at 203,59 size 19x15; Text 'Min'
   IOField "I/O field_2" at 225,75 size 26x19; FormatPattern 999
      ProcessValue <- "Data_DTLData_DTL_Mesin Run[4].SECOND"
   IOField "I/O field_3" at 200,75 size 25x19; FormatPattern 999
      ProcessValue <- "Data_DTLData_DTL_Mesin Run[4].MINUTE"
   TextField "Text field_3" at 30,58 size 144x17; Text 'Time Counter Machine'
   TextField "Text field_4" at 29,75 size 145x19; Text 'Running'
   TextField "Text field_5" at 29,130 size 145x20; Text 'Error'
   IOField "I/O field_24" at 175,75 size 25x19; FormatPattern 999
      ProcessValue <- "Data_DTLData_DTL_Mesin Run[4].HOUR"
   TextField "Text field_13" at 196,74 size 8x17; Text ':'
   TextField "Text field_14" at 196,129 size 8x17; Text ':'
   TextField "Text field_17" at 220,74 size 8x17; Text ':'
   TextField "Text field_18" at 220,129 size 8x17; Text ':'
   TextField "Text field_23" at 196,91 size 8x17; Text ':'
   TextField "Text field_24" at 220,91 size 8x17; Text ':'
   TextField "Text field_26" at 196,109 size 8x17; Text ':'
   TextField "Text field_27" at 220,109 size 8x17; Text ':'
   Button "Button_1" at 47,206 size 90x32; TextOff 'Back To Statistika Data'; TextOn 'Statistika Data'
      on Click: ActivateScreen("Data Statistika", 0)
   Button "Button_3" at 1,205 size 41x34; TextOff 'Main Page'; PictureOff "Home"
      on Click: ActivateScreen("Main Page", 0)
   Button "Button_2" at 236,207 size 80x30; TextOff 'Next Data --->'; TextOn 'Detail Error'
      on Click: ActivateScreen("Error Counter_4", 0)
   Button "Button_4" at 146,207 size 87x30; TextOff '<--- Back Data'; TextOn 'Sloft Data'
      on Click: ActivateScreen("Data Current Shift_4", 0)
   TextField "Text field_1" at 47,0 size 230x18; Text 'CURRENT SHIFT MINUS 4 (Time Data)'

screen "Data Time Current Shift_5" 320x240
   IOField "I/O field_12" at 252,92 size 56x19; FormatPattern 999.99; Unit   %
      ProcessValue <- "Data_Real_%Mesin Run Baypass[5]"
   IOField "I/O field_13" at 252,110 size 56x21; FormatPattern 999.99; Unit   %
      ProcessValue <- "Data_Real_%Mesin Stop[5]"
   IOField "I/O field_14" at 252,130 size 56x20; FormatPattern 999.99; Unit   %
      ProcessValue <- "Data_Real_%Mesin Error[5]"
   IOField "I/O field_11" at 252,75 size 56x18; FormatPattern 999.99; Unit   %
      ProcessValue <- "Data_Real_%Mesin Run[5]"
   IOField "I/O field_6" at 7,24 size 132x18; FormatPattern 9999999999999999999999999999999999999999
      ProcessValue <- "DB_DTL1_Cur_ShiftA_5"
   TextField "Text field_9" at 145,23 size 19x15; Text 'S/D'
   IOField "I/O field_7" at 170,24 size 132x18; FormatPattern 9999999999999999999999999999999999999999
      ProcessValue <- "DB_DTL1_Cur_ShiftB_5"
   TextField "Text field_32" at 7,130 size 21x19; Text '4'
   TextField "Text field_31" at 7,111 size 21x19; Text '3'
   TextField "Text field_30" at 7,92 size 21x19; Text '2'
   TextField "Text field_29" at 7,74 size 21x19; Text '1'
   TextField "Text field_28" at 7,56 size 21x19; Text 'No'
   IOField "I/O field_21" at 225,110 size 26x19; FormatPattern 999
      ProcessValue <- "Data_DTLData_DTL_Mesin Stop[5].SECOND"
   IOField "I/O field_22" at 200,110 size 25x19; FormatPattern 999
      ProcessValue <- "Data_DTLData_DTL_Mesin Stop[5].MINUTE"
   IOField "I/O field_23" at 175,110 size 25x19; FormatPattern 999
      ProcessValue <- "Data_DTLData_DTL_Mesin Stop[5].HOUR"
   TextField "Text field_25" at 29,111 size 145x19; Text 'Stop'
   IOField "I/O field_18" at 225,92 size 26x19; FormatPattern 999
      ProcessValue <- "Data_DTLData_DTL_Mesin Run Baypass[5].SECOND"
   IOField "I/O field_19" at 200,92 size 25x19; FormatPattern 999
      ProcessValue <- "Data_DTLData_DTL_Mesin Run Baypass[5].MINUTE"
   IOField "I/O field_20" at 175,92 size 25x19; FormatPattern 999
      ProcessValue <- "Data_DTLData_DTL_Mesin Run Baypass[5].HOUR"
   TextField "Text field_22" at 29,92 size 145x19; Text 'Running Bypass Stamp'
   TextField "Text field_2" at 176,59 size 24x15; Text 'Hour'
   IOField "I/O field_4" at 225,130 size 26x19; FormatPattern 999
      ProcessValue <- "Data_DTLData_DTL_Mesin Error[5].SECOND"
   IOField "I/O field_5" at 200,130 size 25x19; FormatPattern 999
      ProcessValue <- "Data_DTLData_DTL_Mesin Error[5].MINUTE"
   IOField "I/O field_9" at 175,130 size 25x19; FormatPattern 999
      ProcessValue <- "Data_DTLData_DTL_Mesin Error[5].HOUR"
   TextField "Text field_12" at 229,59 size 19x15; Text 'Sec'
   TextField "Text field_11" at 203,59 size 19x15; Text 'Min'
   IOField "I/O field_2" at 225,75 size 26x19; FormatPattern 999
      ProcessValue <- "Data_DTLData_DTL_Mesin Run[5].SECOND"
   IOField "I/O field_3" at 200,75 size 25x19; FormatPattern 999
      ProcessValue <- "Data_DTLData_DTL_Mesin Run[5].MINUTE"
   TextField "Text field_3" at 30,58 size 144x17; Text 'Time Counter Machine'
   TextField "Text field_4" at 29,75 size 145x19; Text 'Running'
   TextField "Text field_5" at 29,130 size 145x20; Text 'Error'
   IOField "I/O field_24" at 175,75 size 25x19; FormatPattern 999
      ProcessValue <- "Data_DTLData_DTL_Mesin Run[5].HOUR"
   TextField "Text field_13" at 196,74 size 8x17; Text ':'
   TextField "Text field_14" at 196,129 size 8x17; Text ':'
   TextField "Text field_17" at 220,74 size 8x17; Text ':'
   TextField "Text field_18" at 220,129 size 8x17; Text ':'
   TextField "Text field_23" at 196,91 size 8x17; Text ':'
   TextField "Text field_24" at 220,91 size 8x17; Text ':'
   TextField "Text field_26" at 196,109 size 8x17; Text ':'
   TextField "Text field_27" at 220,109 size 8x17; Text ':'
   Button "Button_1" at 47,206 size 90x32; TextOff 'Back To Statistika Data'; TextOn 'Statistika Data'
      on Click: ActivateScreen("Data Statistika", 0)
   Button "Button_3" at 1,205 size 41x34; TextOff 'Main Page'; PictureOff "Home"
      on Click: ActivateScreen("Main Page", 0)
   Button "Button_2" at 236,207 size 80x30; TextOff 'Next Data --->'; TextOn 'Detail Error'
      on Click: ActivateScreen("Error Counter_5", 0)
   Button "Button_4" at 146,207 size 87x30; TextOff '<--- Back Data'; TextOn 'Sloft Data'
      on Click: ActivateScreen("Data Current Shift_5", 0)
   TextField "Text field_1" at 47,0 size 230x18; Text 'CURRENT SHIFT MINUS 5 (Time Data)'
*)